(* Logix 5000 project; controller UOWHF Emulate 5570 rev 30.12; software revision 30.00; part 11 of 13 *)
(* tags used below, declared in another part *)
   UOWHF_Add_c : DINT;
   UOWHF_Msg : DINT[16];
   UOWHF_Result : DINT[16];
(* MainProgram, continued *)

   		UOWHF_Add_c.2:=UOWHF_Result[2].31;
   		UOWHF_Result[2].31:=0;
   		UOWHF_Result[3]:=UOWHF_Result[3] + 1591004397+UOWHF_Add_c;
   		UOWHF_Add_c.3:=UOWHF_Result[3].31;
   		UOWHF_Result[3].31:=0;
   		UOWHF_Result[4]:=UOWHF_Result[4] + 1640170804+UOWHF_Add_c;
   		UOWHF_Add_c.4:=UOWHF_Result[4].31;
   		UOWHF_Result[4].31:=0;
   		UOWHF_Result[5]:=UOWHF_Result[5] + 417190836+UOWHF_Add_c;
   		UOWHF_Add_c.5:=UOWHF_Result[5].31;
   		UOWHF_Result[5].31:=0;
   		UOWHF_Result[6]:=UOWHF_Result[6] + 1926019562+UOWHF_Add_c;
   		UOWHF_Add_c.6:=UOWHF_Result[6].31;
   		UOWHF_Result[6].31:=0;
   		UOWHF_Result[7]:=UOWHF_Result[7] + 695957955+UOWHF_Add_c;
   		UOWHF_Add_c.7:=UOWHF_Result[7].31;
   		UOWHF_Result[7].31:=0;
   		UOWHF_Result[8]:=UOWHF_Result[8] + 1059440084+UOWHF_Add_c;
   		UOWHF_Add_c.8:=UOWHF_Result[8].31;
   		UOWHF_Result[8].31:=0;
   	End_If;
   	If UOWHF_Msg[10].[4] Then
   		UOWHF_Result[0]:=UOWHF_Result[0] + 901796020+UOWHF_Add_c;
   		UOWHF_Add_c.0:=UOWHF_Result[0].31;
   		UOWHF_Result[0].31:=0;
   		UOWHF_Result[1]:=UOWHF_Result[1] + 1127200049+UOWHF_Add_c;
   		UOWHF_Add_c.1:=UOWHF_Result[1].31;
   		UOWHF_Result[1].31:=0;
   		UOWHF_Result[2]:=UOWHF_Result[2] + 1602413067+UOWHF_Add_c;
   		UOWHF_Add_c.2:=UOWHF_Result[2].31;
   		UOWHF_Result[2].31:=0;
   		UOWHF_Result[3]:=UOWHF_Result[3] + 1255033930+UOWHF_Add_c;
   		UOWHF_Add_c.3:=UOWHF_Result[3].31;
   		UOWHF_Result[3].31:=0;
   		UOWHF_Result[4]:=UOWHF_Result[4] + 2144327764+UOWHF_Add_c;
   		UOWHF_Add_c.4:=UOWHF_Result[4].31;
   		UOWHF_Result[4].31:=0;
   		UOWHF_Result[5]:=UOWHF_Result[5] + 1452466792+UOWHF_Add_c;
   		UOWHF_Add_c.5:=UOWHF_Result[5].31;
   		UOWHF_Result[5].31:=0;
   		UOWHF_Result[6]:=UOWHF_Result[6] + 154742090+UOWHF_Add_c;
   		UOWHF_Add_c.6:=UOWHF_Result[6].31;
   		UOWHF_Result[6].31:=0;
   		UOWHF_Result[7]:=UOWHF_Result[7] + 1902468370+UOWHF_Add_c;
   		UOWHF_Add_c.7:=UOWHF_Result[7].31;
   		UOWHF_Result[7].31:=0;
   		UOWHF_Result[8]:=UOWHF_Result[8] + 342884653+UOWHF_Add_c;
   		UOWHF_Add_c.8:=UOWHF_Result[8].31;
   		UOWHF_Result[8].31:=0;
   	End_If;
   	If UOWHF_Msg[10].[5] Then
   		UOWHF_Result[0]:=UOWHF_Result[0] + 868277617+UOWHF_Add_c;
   		UOWHF_Add_c.0:=UOWHF_Result[0].31;
   		UOWHF_Result[0].31:=0;
   		UOWHF_Result[1]:=UOWHF_Result[1] + 1436615864+UOWHF_Add_c;
   		UOWHF_Add_c.1:=UOWHF_Result[1].31;
   		UOWHF_Result[1].31:=0;
   		UOWHF_Result[2]:=UOWHF_Result[2] + 1784814025+UOWHF_Add_c;
   		UOWHF_Add_c.2:=UOWHF_Result[2].31;
   		UOWHF_Result[2].31:=0;
   		UOWHF_Result[3]:=UOWHF_Result[3] + 1380127603+UOWHF_Add_c;
   		UOWHF_Add_c.3:=UOWHF_Result[3].31;
   		UOWHF_Result[3].31:=0;
   		UOWHF_Result[4]:=UOWHF_Result[4] + 1271855125+UOWHF_Add_c;
   		UOWHF_Add_c.4:=UOWHF_Result[4].31;
   		UOWHF_Result[4].31:=0;
   		UOWHF_Result[5]:=UOWHF_Result[5] + 1937374017+UOWHF_Add_c;
   		UOWHF_Add_c.5:=UOWHF_Result[5].31;
   		UOWHF_Result[5].31:=0;
   		UOWHF_Result[6]:=UOWHF_Result[6] + 1845918423+UOWHF_Add_c;
   		UOWHF_Add_c.6:=UOWHF_Result[6].31;
   		UOWHF_Result[6].31:=0;
   		UOWHF_Result[7]:=UOWHF_Result[7] + 1463581006+UOWHF_Add_c;
   		UOWHF_Add_c.7:=UOWHF_Result[7].31;
   		UOWHF_Result[7].31:=0;
   		UOWHF_Result[8]:=UOWHF_Result[8] + 350086967+UOWHF_Add_c;
   		UOWHF_Add_c.8:=UOWHF_Result[8].31;
   		UOWHF_Result[8].31:=0;
   	End_If;
   	If UOWHF_Msg[10].[6] Then
   		UOWHF_Result[0]:=UOWHF_Result[0] + 1588271974+UOWHF_Add_c;
   		UOWHF_Add_c.0:=UOWHF_Result[0].31;
   		UOWHF_Result[0].31:=0;
   		UOWHF_Result[1]:=UOWHF_Result[1] + 586756377+UOWHF_Add_c;
   		UOWHF_Add_c.1:=UOWHF_Result[1].31;
   		UOWHF_Result[1].31:=0;
   		UOWHF_Result[2]:=UOWHF_Result[2] + 559516102+UOWHF_Add_c;
   		UOWHF_Add_c.2:=UOWHF_Result[2].31;
   		UOWHF_Result[2].31:=0;
   		UOWHF_Result[3]:=UOWHF_Result[3] + 331741523+UOWHF_Add_c;
   		UOWHF_Add_c.3:=UOWHF_Result[3].31;
   		UOWHF_Result[3].31:=0;
   		UOWHF_Result[4]:=UOWHF_Result[4] + 1880781678+UOWHF_Add_c;
   		UOWHF_Add_c.4:=UOWHF_Result[4].31;
   		UOWHF_Result[4].31:=0;
   		UOWHF_Result[5]:=UOWHF_Result[5] + 1152892566+UOWHF_Add_c;
   		UOWHF_Add_c.5:=UOWHF_Result[5].31;
   		UOWHF_Result[5].31:=0;
   		UOWHF_Result[6]:=UOWHF_Result[6] + 2047233698+UOWHF_Add_c;
   		UOWHF_Add_c.6:=UOWHF_Result[6].31;
   		UOWHF_Result[6].31:=0;
   		UOWHF_Result[7]:=UOWHF_Result[7] + 1642594289+UOWHF_Add_c;
   		UOWHF_Add_c.7:=UOWHF_Result[7].31;
   		UOWHF_Result[7].31:=0;
   		UOWHF_Result[8]:=UOWHF_Result[8] + 376585573+UOWHF_Add_c;
   		UOWHF_Add_c.8:=UOWHF_Result[8].31;
   		UOWHF_Result[8].31:=0;
   	End_If;
   	If UOWHF_Msg[10].[7] Then
   		UOWHF_Result[0]:=UOWHF_Result[0] + 1020715491+UOWHF_Add_c;
   		UOWHF_Add_c.0:=UOWHF_Result[0].31;
   		UOWHF_Result[0].31:=0;
   		UOWHF_Result[1]:=UOWHF_Result[1] + 1857205629+UOWHF_Add_c;
   		UOWHF_Add_c.1:=UOWHF_Result[1].31;
   		UOWHF_Result[1].31:=0;
   		UOWHF_Result[2]:=UOWHF_Result[2] + 16853309+UOWHF_Add_c;
   		UOWHF_Add_c.2:=UOWHF_Result[2].31;
   		UOWHF_Result[2].31:=0;
   		UOWHF_Result[3]:=UOWHF_Result[3] + 1231994168+UOWHF_Add_c;
   		UOWHF_Add_c.3:=UOWHF_Result[3].31;
   		UOWHF_Result[3].31:=0;
   		UOWHF_Result[4]:=UOWHF_Result[4] + 423998966+UOWHF_Add_c;
   		UOWHF_Add_c.4:=UOWHF_Result[4].31;
   		UOWHF_Result[4].31:=0;
   		UOWHF_Result[5]:=UOWHF_Result[5] + 1299862752+UOWHF_Add_c;
   		UOWHF_Add_c.5:=UOWHF_Result[5].31;
   		UOWHF_Result[5].31:=0;
   		UOWHF_Result[6]:=UOWHF_Result[6] + 652509862+UOWHF_Add_c;
   		UOWHF_Add_c.6:=UOWHF_Result[6].31;
   		UOWHF_Result[6].31:=0;
   		UOWHF_Result[7]:=UOWHF_Result[7] + 15353685+UOWHF_Add_c;
   		UOWHF_Add_c.7:=UOWHF_Result[7].31;
   		UOWHF_Result[7].31:=0;
   		UOWHF_Result[8]:=UOWHF_Result[8] + 2001428660+UOWHF_Add_c;
   		UOWHF_Add_c.8:=UOWHF_Result[8].31;
   		UOWHF_Result[8].31:=0;
   	End_If;
   	If UOWHF_Msg[10].[8] Then
   		UOWHF_Result[0]:=UOWHF_Result[0] + 813810484+UOWHF_Add_c;
   		UOWHF_Add_c.0:=UOWHF_Result[0].31;
   		UOWHF_Result[0].31:=0;
   		UOWHF_Result[1]:=UOWHF_Result[1] + 1003989381+UOWHF_Add_c;
   		UOWHF_Add_c.1:=UOWHF_Result[1].31;
   		UOWHF_Result[1].31:=0;
   		UOWHF_Result[2]:=UOWHF_Result[2] + 738018774+UOWHF_Add_c;
   		UOWHF_Add_c.2:=UOWHF_Result[2].31;
   		UOWHF_Result[2].31:=0;
   		UOWHF_Result[3]:=UOWHF_Result[3] + 443461312+UOWHF_Add_c;
   		UOWHF_Add_c.3:=UOWHF_Result[3].31;
   		UOWHF_Result[3].31:=0;
   		UOWHF_Result[4]:=UOWHF_Result[4] + 1637414295+UOWHF_Add_c;
   		UOWHF_Add_c.4:=UOWHF_Result[4].31;
   		UOWHF_Result[4].31:=0;
   		UOWHF_Result[5]:=UOWHF_Result[5] + 157939787+UOWHF_Add_c;
   		UOWHF_Add_c.5:=UOWHF_Result[5].31;
   		UOWHF_Result[5].31:=0;
   		UOWHF_Result[6]:=UOWHF_Result[6] + 712235666+UOWHF_Add_c;
   		UOWHF_Add_c.6:=UOWHF_Result[6].31;
   		UOWHF_Result[6].31:=0;
   		UOWHF_Result[7]:=UOWHF_Result[7] + 1688386276+UOWHF_Add_c;
   		UOWHF_Add_c.7:=UOWHF_Result[7].31;
   		UOWHF_Result[7].31:=0;
   		UOWHF_Result[8]:=UOWHF_Result[8] + 2013177678+UOWHF_Add_c;
   		UOWHF_Add_c.8:=UOWHF_Result[8].31;
   		UOWHF_Result[8].31:=0;
   	End_If;
   	If UOWHF_Msg[10].[9] Then
   		UOWHF_Result[0]:=UOWHF_Result[0] + 1535414445+UOWHF_Add_c;
   		UOWHF_Add_c.0:=UOWHF_Result[0].31;
   		UOWHF_Result[0].31:=0;
   		UOWHF_Result[1]:=UOWHF_Result[1] + 1615623515+UOWHF_Add_c;
   		UOWHF_Add_c.1:=UOWHF_Result[1].31;
   		UOWHF_Result[1].31:=0;
   		UOWHF_Result[2]:=UOWHF_Result[2] + 1360597756+UOWHF_Add_c;
   		UOWHF_Add_c.2:=UOWHF_Result[2].31;
   		UOWHF_Result[2].31:=0;
   		UOWHF_Result[3]:=UOWHF_Result[3] + 1573823097+UOWHF_Add_c;
   		UOWHF_Add_c.3:=UOWHF_Result[3].31;
   		UOWHF_Result[3].31:=0;
   		UOWHF_Result[4]:=UOWHF_Result[4] + 1281710714+UOWHF_Add_c;
   		UOWHF_Add_c.4:=UOWHF_Result[4].31;
   		UOWHF_Result[4].31:=0;
   		UOWHF_Result[5]:=UOWHF_Result[5] + 1453733315+UOWHF_Add_c;
   		UOWHF_Add_c.5:=UOWHF_Result[5].31;
   		UOWHF_Result[5].31:=0;
   		UOWHF_Result[6]:=UOWHF_Result[6] + 369997754+UOWHF_Add_c;
   		UOWHF_Add_c.6:=UOWHF_Result[6].31;
   		UOWHF_Result[6].31:=0;
   		UOWHF_Result[7]:=UOWHF_Result[7] + 1856281529+UOWHF_Add_c;
   		UOWHF_Add_c.7:=UOWHF_Result[7].31;
   		UOWHF_Result[7].31:=0;
   		UOWHF_Result[8]:=UOWHF_Result[8] + 1847238559+UOWHF_Add_c;
   		UOWHF_Add_c.8:=UOWHF_Result[8].31;
   		UOWHF_Result[8].31:=0;
   	End_If;
   	If UOWHF_Msg[10].[10] Then
   		UOWHF_Result[0]:=UOWHF_Result[0] + 1061749827+UOWHF_Add_c;
   		UOWHF_Add_c.0:=UOWHF_Result[0].31;
   		UOWHF_Result[0].31:=0;
   		UOWHF_Result[1]:=UOWHF_Result[1] + 842932244+UOWHF_Add_c;
   		UOWHF_Add_c.1:=UOWHF_Result[1].31;
   		UOWHF_Result[1].31:=0;
   		UOWHF_Result[2]:=UOWHF_Result[2] + 1033461891+UOWHF_Add_c;
   		UOWHF_Add_c.2:=UOWHF_Result[2].31;
   		UOWHF_Result[2].31:=0;
   		UOWHF_Result[3]:=UOWHF_Result[3] + 379746348+UOWHF_Add_c;
   		UOWHF_Add_c.3:=UOWHF_Result[3].31;
   		UOWHF_Result[3].31:=0;
   		UOWHF_Result[4]:=UOWHF_Result[4] + 685495130+UOWHF_Add_c;
   		UOWHF_Add_c.4:=UOWHF_Result[4].31;
   		UOWHF_Result[4].31:=0;
   		UOWHF_Result[5]:=UOWHF_Result[5] + 958802377+UOWHF_Add_c;
   		UOWHF_Add_c.5:=UOWHF_Result[5].31;
   		UOWHF_Result[5].31:=0;
   		UOWHF_Result[6]:=UOWHF_Result[6] + 129067151+UOWHF_Add_c;
   		UOWHF_Add_c.6:=UOWHF_Result[6].31;
   		UOWHF_Result[6].31:=0;
   		UOWHF_Result[7]:=UOWHF_Result[7] + 1694766568+UOWHF_Add_c;
   		UOWHF_Add_c.7:=UOWHF_Result[7].31;
   		UOWHF_Result[7].31:=0;
   		UOWHF_Result[8]:=UOWHF_Result[8] + 1431412769+UOWHF_Add_c;
   		UOWHF_Add_c.8:=UOWHF_Result[8].31;
   		UOWHF_Result[8].31:=0;
   	End_If;
   	If UOWHF_Msg[10].[11] Then
   		UOWHF_Result[0]:=UOWHF_Result[0] + 1646350318+UOWHF_Add_c;
   		UOWHF_Add_c.0:=UOWHF_Result[0].31;
   		UOWHF_Result[0].31:=0;
   		UOWHF_Result[1]:=UOWHF_Result[1] + 1974652699+UOWHF_Add_c;
   		UOWHF_Add_c.1:=UOWHF_Result[1].31;
   		UOWHF_Result[1].31:=0;
   		UOWHF_Result[2]:=UOWHF_Result[2] + 325775484+UOWHF_Add_c;
   		UOWHF_Add_c.2:=UOWHF_Result[2].31;
   		UOWHF_Result[2].31:=0;
   		UOWHF_Result[3]:=UOWHF_Result[3] + 83362006+UOWHF_Add_c;
   		UOWHF_Add_c.3:=UOWHF_Result[3].31;
   		UOWHF_Result[3].31:=0;
   		UOWHF_Result[4]:=UOWHF_Result[4] + 262049431+UOWHF_Add_c;
   		UOWHF_Add_c.4:=UOWHF_Result[4].31;
   		UOWHF_Result[4].31:=0;
   		UOWHF_Result[5]:=UOWHF_Result[5] + 1644755762+UOWHF_Add_c;
   		UOWHF_Add_c.5:=UOWHF_Result[5].31;
   		UOWHF_Result[5].31:=0;
   		UOWHF_Result[6]:=UOWHF_Result[6] + 790241358+UOWHF_Add_c;
   		UOWHF_Add_c.6:=UOWHF_Result[6].31;
   		UOWHF_Result[6].31:=0;
   		UOWHF_Result[7]:=UOWHF_Result[7] + 2126439262+UOWHF_Add_c;
   		UOWHF_Add_c.7:=UOWHF_Result[7].31;
   		UOWHF_Result[7].31:=0;
   		UOWHF_Result[8]:=UOWHF_Result[8] + 1052212769+UOWHF_Add_c;
   		UOWHF_Add_c.8:=UOWHF_Result[8].31;
   		UOWHF_Result[8].31:=0;
   	End_If;
   	If UOWHF_Msg[10].[12] Then
   		UOWHF_Result[0]:=UOWHF_Result[0] + 955937059+UOWHF_Add_c;
   		UOWHF_Add_c.0:=UOWHF_Result[0].31;
   		UOWHF_Result[0].31:=0;
   		UOWHF_Result[1]:=UOWHF_Result[1] + 936365642+UOWHF_Add_c;
   		UOWHF_Add_c.1:=UOWHF_Result[1].31;
   		UOWHF_Result[1].31:=0;
   		UOWHF_Result[2]:=UOWHF_Result[2] + 498042732+UOWHF_Add_c;
   		UOWHF_Add_c.2:=UOWHF_Result[2].31;
   		UOWHF_Result[2].31:=0;
   		UOWHF_Result[3]:=UOWHF_Result[3] + 238009702+UOWHF_Add_c;
   		UOWHF_Add_c.3:=UOWHF_Result[3].31;
   		UOWHF_Result[3].31:=0;
   		UOWHF_Result[4]:=UOWHF_Result[4] + 36957456+UOWHF_Add_c;
   		UOWHF_Add_c.4:=UOWHF_Result[4].31;
   		UOWHF_Result[4].31:=0;
   		UOWHF_Result[5]:=UOWHF_Result[5] + 598813011+UOWHF_Add_c;
   		UOWHF_Add_c.5:=UOWHF_Result[5].31;
   		UOWHF_Result[5].31:=0;
   		UOWHF_Result[6]:=UOWHF_Result[6] + 426350274+UOWHF_Add_c;
   		UOWHF_Add_c.6:=UOWHF_Result[6].31;
   		UOWHF_Result[6].31:=0;
   		UOWHF_Result[7]:=UOWHF_Result[7] + 102852187+UOWHF_Add_c;
   		UOWHF_Add_c.7:=UOWHF_Result[7].31;
   		UOWHF_Result[7].31:=0;
   		UOWHF_Result[8]:=UOWHF_Result[8] + 1154127904+UOWHF_Add_c;
   		UOWHF_Add_c.8:=UOWHF_Result[8].31;
   		UOWHF_Result[8].31:=0;
   	End_If;
   	If UOWHF_Msg[10].[13] Then
   		UOWHF_Result[0]:=UOWHF_Result[0] + 1268816444+UOWHF_Add_c;
   		UOWHF_Add_c.0:=UOWHF_Result[0].31;
   		UOWHF_Result[0].31:=0;
   		UOWHF_Result[1]:=UOWHF_Result[1] + 1033144398+UOWHF_Add_c;
   		UOWHF_Add_c.1:=UOWHF_Result[1].31;
   		UOWHF_Result[1].31:=0;
   		UOWHF_Result[2]:=UOWHF_Result[2] + 2027448386+UOWHF_Add_c;
   		UOWHF_Add_c.2:=UOWHF_Result[2].31;
   		UOWHF_Result[2].31:=0;
   		UOWHF_Result[3]:=UOWHF_Result[3] + 885764043+UOWHF_Add_c;
   		UOWHF_Add_c.3:=UOWHF_Result[3].31;
   		UOWHF_Result[3].31:=0;
   		UOWHF_Result[4]:=UOWHF_Result[4] + 1657422268+UOWHF_Add_c;
   		UOWHF_Add_c.4:=UOWHF_Result[4].31;
   		UOWHF_Result[4].31:=0;
   		UOWHF_Result[5]:=UOWHF_Result[5] + 1988850223+UOWHF_Add_c;
   		UOWHF_Add_c.5:=UOWHF_Result[5].31;
   		UOWHF_Result[5].31:=0;
   		UOWHF_Result[6]:=UOWHF_Result[6] + 1530930092+UOWHF_Add_c;
   		UOWHF_Add_c.6:=UOWHF_Result[6].31;
   		UOWHF_Result[6].31:=0;
   		UOWHF_Result[7]:=UOWHF_Result[7] + 2006297248+UOWHF_Add_c;
   		UOWHF_Add_c.7:=UOWHF_Result[7].31;
   		UOWHF_Result[7].31:=0;
   		UOWHF_Result[8]:=UOWHF_Result[8] + 2077959681+UOWHF_Add_c;
   		UOWHF_Add_c.8:=UOWHF_Result[8].31;
   		UOWHF_Result[8].31:=0;
   	End_If;
   	If UOWHF_Msg[10].[14] Then
   		UOWHF_Result[0]:=UOWHF_Result[0] + 1110917864+UOWHF_Add_c;
   		UOWHF_Add_c.0:=UOWHF_Result[0].31;
   		UOWHF_Result[0].31:=0;
   		UOWHF_Result[1]:=UOWHF_Result[1] + 1451124381+UOWHF_Add_c;
   		UOWHF_Add_c.1:=UOWHF_Result[1].31;
   		UOWHF_Result[1].31:=0;
   		UOWHF_Result[2]:=UOWHF_Result[2] + 1354761017+UOWHF_Add_c;
   		UOWHF_Add_c.2:=UOWHF_Result[2].31;
   		UOWHF_Result[2].31:=0;
   		UOWHF_Result[3]:=UOWHF_Result[3] + 38190742+UOWHF_Add_c;
   		UOWHF_Add_c.3:=UOWHF_Result[3].31;
   		UOWHF_Result[3].31:=0;
   		UOWHF_Result[4]:=UOWHF_Result[4] + 1921805953+UOWHF_Add_c;
   		UOWHF_Add_c.4:=UOWHF_Result[4].31;
   		UOWHF_Result[4].31:=0;
   		UOWHF_Result[5]:=UOWHF_Result[5] + 1941105002+UOWHF_Add_c;
   		UOWHF_Add_c.5:=UOWHF_Result[5].31;
   		UOWHF_Result[5].31:=0;
   		UOWHF_Result[6]:=UOWHF_Result[6] + 1703548468+UOWHF_Add_c;
   		UOWHF_Add_c.6:=UOWHF_Result[6].31;
   		UOWHF_Result[6].31:=0;
   		UOWHF_Result[7]:=UOWHF_Result[7] + 186991094+UOWHF_Add_c;
   		UOWHF_Add_c.7:=UOWHF_Result[7].31;
   		UOWHF_Result[7].31:=0;
   		UOWHF_Result[8]:=UOWHF_Result[8] + 714064657+UOWHF_Add_c;
   		UOWHF_Add_c.8:=UOWHF_Result[8].31;
   		UOWHF_Result[8].31:=0;
   	End_If;
   	If UOWHF_Msg[10].[15] Then
   		UOWHF_Result[0]:=UOWHF_Result[0] + 1961147110+UOWHF_Add_c;
   		UOWHF_Add_c.0:=UOWHF_Result[0].31;
   		UOWHF_Result[0].31:=0;
   		UOWHF_Result[1]:=UOWHF_Result[1] + 12565547+UOWHF_Add_c;
   		UOWHF_Add_c.1:=UOWHF_Result[1].31;
   		UOWHF_Result[1].31:=0;
   		UOWHF_Result[2]:=UOWHF_Result[2] + 567043951+UOWHF_Add_c;
   		UOWHF_Add_c.2:=UOWHF_Result[2].31;
   		UOWHF_Result[2].31:=0;
   		UOWHF_Result[3]:=UOWHF_Result[3] + 65949662+UOWHF_Add_c;
   		UOWHF_Add_c.3:=UOWHF_Result[3].31;
   		UOWHF_Result[3].31:=0;
   		UOWHF_Result[4]:=UOWHF_Result[4] + 1646539206+UOWHF_Add_c;
   		UOWHF_Add_c.4:=UOWHF_Result[4].31;
   		UOWHF_Result[4].31:=0;
   		UOWHF_Result[5]:=UOWHF_Result[5] + 1708716662+UOWHF_Add_c;
   		UOWHF_Add_c.5:=UOWHF_Result[5].31;
   		UOWHF_Result[5].31:=0;
   		UOWHF_Result[6]:=UOWHF_Result[6] + 1848936862+UOWHF_Add_c;
   		UOWHF_Add_c.6:=UOWHF_Result[6].31;
   		UOWHF_Result[6].31:=0;
   		UOWHF_Result[7]:=UOWHF_Result[7] + 1900654345+UOWHF_Add_c;
   		UOWHF_Add_c.7:=UOWHF_Result[7].31;
   		UOWHF_Result[7].31:=0;
   		UOWHF_Result[8]:=UOWHF_Result[8] + 1004361316+UOWHF_Add_c;
   		UOWHF_Add_c.8:=UOWHF_Result[8].31;
   		UOWHF_Result[8].31:=0;
   	End_If;
   	If UOWHF_Msg[10].[16] Then
   		UOWHF_Result[0]:=UOWHF_Result[0] + 415520432+UOWHF_Add_c;
   		UOWHF_Add_c.0:=UOWHF_Result[0].31;
   		UOWHF_Result[0].31:=0;
   		UOWHF_Result[1]:=UOWHF_Result[1] + 351467464+UOWHF_Add_c;
   		UOWHF_Add_c.1:=UOWHF_Result[1].31;
   		UOWHF_Result[1].31:=0;
   		UOWHF_Result[2]:=UOWHF_Result[2] + 654166220+UOWHF_Add_c;
   		UOWHF_Add_c.2:=UOWHF_Result[2].31;
   		UOWHF_Result[2].31:=0;
   		UOWHF_Result[3]:=UOWHF_Result[3] + 741029837+UOWHF_Add_c;
   		UOWHF_Add_c.3:=UOWHF_Result[3].31;
   		UOWHF_Result[3].31:=0;
   		UOWHF_Result[4]:=UOWHF_Result[4] + 1981690344+UOWHF_Add_c;
   		UOWHF_Add_c.4:=UOWHF_Result[4].31;
   		UOWHF_Result[4].31:=0;
   		UOWHF_Result[5]:=UOWHF_Result[5] + 19210638+UOWHF_Add_c;
   		UOWHF_Add_c.5:=UOWHF_Result[5].31;
   		UOWHF_Result[5].31:=0;
   		UOWHF_Result[6]:=UOWHF_Result[6] + 566229794+UOWHF_Add_c;
   		UOWHF_Add_c.6:=UOWHF_Result[6].31;
   		UOWHF_Result[6].31:=0;
   		UOWHF_Result[7]:=UOWHF_Result[7] + 625793338+UOWHF_Add_c;
   		UOWHF_Add_c.7:=UOWHF_Result[7].31;
   		UOWHF_Result[7].31:=0;
   		UOWHF_Result[8]:=UOWHF_Result[8] + 386405378+UOWHF_Add_c;
   		UOWHF_Add_c.8:=UOWHF_Result[8].31;
   		UOWHF_Result[8].31:=0;
   	End_If;
   	If UOWHF_Msg[10].[17] Then
   		UOWHF_Result[0]:=UOWHF_Result[0] + 1499883797+UOWHF_Add_c;
   		UOWHF_Add_c.0:=UOWHF_Result[0].31;
   		UOWHF_Result[0].31:=0;
   		UOWHF_Result[1]:=UOWHF_Result[1] + 129680376+UOWHF_Add_c;
   		UOWHF_Add_c.1:=UOWHF_Result[1].31;
   		UOWHF_Result[1].31:=0;
   		UOWHF_Result[2]:=UOWHF_Result[2] + 700971919+UOWHF_Add_c;
   		UOWHF_Add_c.2:=UOWHF_Result[2].31;
   		UOWHF_Result[2].31:=0;
   		UOWHF_Result[3]:=UOWHF_Result[3] + 56395807+UOWHF_Add_c;
   		UOWHF_Add_c.3:=UOWHF_Result[3].31;
   		UOWHF_Result[3].31:=0;
   		UOWHF_Result[4]:=UOWHF_Result[4] + 1355965327+UOWHF_Add_c;
   		UOWHF_Add_c.4:=UOWHF_Result[4].31;
   		UOWHF_Result[4].31:=0;
   		UOWHF_Result[5]:=UOWHF_Result[5] + 1408183226+UOWHF_Add_c;
   		UOWHF_Add_c.5:=UOWHF_Result[5].31;
   		UOWHF_Result[5].31:=0;
   		UOWHF_Result[6]:=UOWHF_Result[6] + 2071090026+UOWHF_Add_c;
   		UOWHF_Add_c.6:=UOWHF_Result[6].31;
   		UOWHF_Result[6].31:=0;
   		UOWHF_Result[7]:=UOWHF_Result[7] + 1334749712+UOWHF_Add_c;
   		UOWHF_Add_c.7:=UOWHF_Result[7].31;
   		UOWHF_Result[7].31:=0;
   		UOWHF_Result[8]:=UOWHF_Result[8] + 894206129+UOWHF_Add_c;
   		UOWHF_Add_c.8:=UOWHF_Result[8].31;
   		UOWHF_Result[8].31:=0;
   	End_If;
   	If UOWHF_Msg[10].[18] Then
   		UOWHF_Result[0]:=UOWHF_Result[0] + 611633887+UOWHF_Add_c;
   		UOWHF_Add_c.0:=UOWHF_Result[0].31;
   		UOWHF_Result[0].31:=0;
   		UOWHF_Result[1]:=UOWHF_Result[1] + 220479088+UOWHF_Add_c;
   		UOWHF_Add_c.1:=UOWHF_Result[1].31;
   		UOWHF_Result[1].31:=0;
   		UOWHF_Result[2]:=UOWHF_Result[2] + 774163886+UOWHF_Add_c;
   		UOWHF_Add_c.2:=UOWHF_Result[2].31;
   		UOWHF_Result[2].31:=0;
   		UOWHF_Result[3]:=UOWHF_Result[3] + 244973967+UOWHF_Add_c;
   		UOWHF_Add_c.3:=UOWHF_Result[3].31;
   		UOWHF_Result[3].31:=0;
   		UOWHF_Result[4]:=UOWHF_Result[4] + 906891116+UOWHF_Add_c;
   		UOWHF_Add_c.4:=UOWHF_Result[4].31;
   		UOWHF_Result[4].31:=0;
   		UOWHF_Result[5]:=UOWHF_Result[5] + 2010017338+UOWHF_Add_c;
   		UOWHF_Add_c.5:=UOWHF_Result[5].31;
   		UOWHF_Result[5].31:=0;
   		UOWHF_Result[6]:=UOWHF_Result[6] + 1437360572+UOWHF_Add_c;
   		UOWHF_Add_c.6:=UOWHF_Result[6].31;
   		UOWHF_Result[6].31:=0;
   		UOWHF_Result[7]:=UOWHF_Result[7] + 1208873370+UOWHF_Add_c;
   		UOWHF_Add_c.7:=UOWHF_Result[7].31;
   		UOWHF_Result[7].31:=0;
   		UOWHF_Result[8]:=UOWHF_Result[8] + 73161532+UOWHF_Add_c;
   		UOWHF_Add_c.8:=UOWHF_Result[8].31;
   		UOWHF_Result[8].31:=0;
   	End_If;
   	If UOWHF_Msg[10].[19] Then
   		UOWHF_Result[0]:=UOWHF_Result[0] + 1276434743+UOWHF_Add_c;
   		UOWHF_Add_c.0:=UOWHF_Result[0].31;
   		UOWHF_Result[0].31:=0;
   		UOWHF_Result[1]:=UOWHF_Result[1] + 923954815+UOWHF_Add_c;
   		UOWHF_Add_c.1:=UOWHF_Result[1].31;
   		UOWHF_Result[1].31:=0;
   		UOWHF_Result[2]:=UOWHF_Result[2] + 2127328610+UOWHF_Add_c;
   		UOWHF_Add_c.2:=UOWHF_Result[2].31;
   		UOWHF_Result[2].31:=0;
   		UOWHF_Result[3]:=UOWHF_Result[3] + 1862713612+UOWHF_Add_c;
   		UOWHF_Add_c.3:=UOWHF_Result[3].31;
   		UOWHF_Result[3].31:=0;
   		UOWHF_Result[4]:=UOWHF_Result[4] + 1878938249+UOWHF_Add_c;
   		UOWHF_Add_c.4:=UOWHF_Result[4].31;
   		UOWHF_Result[4].31:=0;
   		UOWHF_Result[5]:=UOWHF_Result[5] + 1189510329+UOWHF_Add_c;
   		UOWHF_Add_c.5:=UOWHF_Result[5].31;
   		UOWHF_Result[5].31:=0;
   		UOWHF_Result[6]:=UOWHF_Result[6] + 1679535384+UOWHF_Add_c;
   		UOWHF_Add_c.6:=UOWHF_Result[6].31;
   		UOWHF_Result[6].31:=0;
   		UOWHF_Result[7]:=UOWHF_Result[7] + 1749990172+UOWHF_Add_c;
   		UOWHF_Add_c.7:=UOWHF_Result[7].31;
   		UOWHF_Result[7].31:=0;
   		UOWHF_Result[8]:=UOWHF_Result[8] + 1880399620+UOWHF_Add_c;
   		UOWHF_Add_c.8:=UOWHF_Result[8].31;
   		UOWHF_Result[8].31:=0;
   	End_If;
   	If UOWHF_Msg[10].[20] Then
   		UOWHF_Result[0]:=UOWHF_Result[0] + 1067539284+UOWHF_Add_c;
   		UOWHF_Add_c.0:=UOWHF_Result[0].31;
   		UOWHF_Result[0].31:=0;
   		UOWHF_Result[1]:=UOWHF_Result[1] + 1218546281+UOWHF_Add_c;
   		UOWHF_Add_c.1:=UOWHF_Result[1].31;
   		UOWHF_Result[1].31:=0;
   		UOWHF_Result[2]:=UOWHF_Result[2] + 1692266167+UOWHF_Add_c;
   		UOWHF_Add_c.2:=UOWHF_Result[2].31;
   		UOWHF_Result[2].31:=0;
   		UOWHF_Result[3]:=UOWHF_Result[3] + 844450602+UOWHF_Add_c;
   		UOWHF_Add_c.3:=UOWHF_Result[3].31;
   		UOWHF_Result[3].31:=0;
   		UOWHF_Result[4]:=UOWHF_Result[4] + 1351238461+UOWHF_Add_c;
   		UOWHF_Add_c.4:=UOWHF_Result[4].31;
   		UOWHF_Result[4].31:=0;
   		UOWHF_Result[5]:=UOWHF_Result[5] + 2074939840+UOWHF_Add_c;
   		UOWHF_Add_c.5:=UOWHF_Result[5].31;
   		UOWHF_Result[5].31:=0;
   		UOWHF_Result[6]:=UOWHF_Result[6] + 54095456+UOWHF_Add_c;
   		UOWHF_Add_c.6:=UOWHF_Result[6].31;
   		UOWHF_Result[6].31:=0;
   		UOWHF_Result[7]:=UOWHF_Result[7] + 1472659390+UOWHF_Add_c;
   		UOWHF_Add_c.7:=UOWHF_Result[7].31;
   		UOWHF_Result[7].31:=0;
   		UOWHF_Result[8]:=UOWHF_Result[8] + 78847011+UOWHF_Add_c;
   		UOWHF_Add_c.8:=UOWHF_Result[8].31;
   		UOWHF_Result[8].31:=0;
   	End_If;
   	If UOWHF_Msg[10].[21] Then
   		UOWHF_Result[0]:=UOWHF_Result[0] + 615459290+UOWHF_Add_c;
   		UOWHF_Add_c.0:=UOWHF_Result[0].31;
   		UOWHF_Result[0].31:=0;
   		UOWHF_Result[1]:=UOWHF_Result[1] + 628300652+UOWHF_Add_c;
   		UOWHF_Add_c.1:=UOWHF_Result[1].31;
   		UOWHF_Result[1].31:=0;
   		UOWHF_Result[2]:=UOWHF_Result[2] + 913630562+UOWHF_Add_c;
   		UOWHF_Add_c.2:=UOWHF_Result[2].31;
   		UOWHF_Result[2].31:=0;
   		UOWHF_Result[3]:=UOWHF_Result[3] + 1573973421+UOWHF_Add_c;
   		UOWHF_Add_c.3:=UOWHF_Result[3].31;
   		UOWHF_Result[3].31:=0;
   		UOWHF_Result[4]:=UOWHF_Result[4] + 842720559+UOWHF_Add_c;
   		UOWHF_Add_c.4:=UOWHF_Result[4].31;
   		UOWHF_Result[4].31:=0;
   		UOWHF_Result[5]:=UOWHF_Result[5] + 1465717949+UOWHF_Add_c;
   		UOWHF_Add_c.5:=UOWHF_Result[5].31;
   		UOWHF_Result[5].31:=0;
   		UOWHF_Result[6]:=UOWHF_Result[6] + 1475649611+UOWHF_Add_c;
   		UOWHF_Add_c.6:=UOWHF_Result[6].31;
   		UOWHF_Result[6].31:=0;
   		UOWHF_Result[7]:=UOWHF_Result[7] + 1123747716+UOWHF_Add_c;
   		UOWHF_Add_c.7:=UOWHF_Result[7].31;
   		UOWHF_Result[7].31:=0;
   		UOWHF_Result[8]:=UOWHF_Result[8] + 593611670+UOWHF_Add_c;
   		UOWHF_Add_c.8:=UOWHF_Result[8].31;
   		UOWHF_Result[8].31:=0;
   	End_If;
   	If UOWHF_Msg[10].[22] Then
   		UOWHF_Result[0]:=UOWHF_Result[0] + 333024015+UOWHF_Add_c;
   		UOWHF_Add_c.0:=UOWHF_Result[0].31;
   		UOWHF_Result[0].31:=0;
   		UOWHF_Result[1]:=UOWHF_Result[1] + 649171931+UOWHF_Add_c;
   		UOWHF_Add_c.1:=UOWHF_Result[1].31;
   		UOWHF_Result[1].31:=0;
   		UOWHF_Result[2]:=UOWHF_Result[2] + 1523497291+UOWHF_Add_c;
   		UOWHF_Add_c.2:=UOWHF_Result[2].31;
   		UOWHF_Result[2].31:=0;
   		UOWHF_Result[3]:=UOWHF_Result[3] + 1354970453+UOWHF_Add_c;
   		UOWHF_Add_c.3:=UOWHF_Result[3].31;
   		UOWHF_Result[3].31:=0;
   		UOWHF_Result[4]:=UOWHF_Result[4] + 72262000+UOWHF_Add_c;
   		UOWHF_Add_c.4:=UOWHF_Result[4].31;
   		UOWHF_Result[4].31:=0;
   		UOWHF_Result[5]:=UOWHF_Result[5] + 246209462+UOWHF_Add_c;
   		UOWHF_Add_c.5:=UOWHF_Result[5].31;
   		UOWHF_Result[5].31:=0;
   		UOWHF_Result[6]:=UOWHF_Result[6] + 1497013496+UOWHF_Add_c;
   		UOWHF_Add_c.6:=UOWHF_Result[6].31;
   		UOWHF_Result[6].31:=0;
   		UOWHF_Result[7]:=UOWHF_Result[7] + 133031163+UOWHF_Add_c;
   		UOWHF_Add_c.7:=UOWHF_Result[7].31;
   		UOWHF_Result[7].31:=0;
   		UOWHF_Result[8]:=UOWHF_Result[8] + 1209415317+UOWHF_Add_c;
   		UOWHF_Add_c.8:=UOWHF_Result[8].31;
   		UOWHF_Result[8].31:=0;
   	End_If;
   	If UOWHF_Msg[10].[23] Then
   		UOWHF_Result[0]:=UOWHF_Result[0] + 1058819959+UOWHF_Add_c;
   		UOWHF_Add_c.0:=UOWHF_Result[0].31;
   		UOWHF_Result[0].31:=0;
   		UOWHF_Result[1]:=UOWHF_Result[1] + 1490152365+UOWHF_Add_c;
   		UOWHF_Add_c.1:=UOWHF_Result[1].31;
   		UOWHF_Result[1].31:=0;
   		UOWHF_Result[2]:=UOWHF_Result[2] + 750844208+UOWHF_Add_c;
   		UOWHF_Add_c.2:=UOWHF_Result[2].31;
   		UOWHF_Result[2].31:=0;
   		UOWHF_Result[3]:=UOWHF_Result[3] + 69060592+UOWHF_Add_c;
   		UOWHF_Add_c.3:=UOWHF_Result[3].31;
   		UOWHF_Result[3].31:=0;
   		UOWHF_Result[4]:=UOWHF_Result[4] + 1239135017+UOWHF_Add_c;
   		UOWHF_Add_c.4:=UOWHF_Result[4].31;
   		UOWHF_Result[4].31:=0;
   		UOWHF_Result[5]:=UOWHF_Result[5] + 1324052255+UOWHF_Add_c;
   		UOWHF_Add_c.5:=UOWHF_Result[5].31;
   		UOWHF_Result[5].31:=0;
   		UOWHF_Result[6]:=UOWHF_Result[6] + 464992231+UOWHF_Add_c;
   		UOWHF_Add_c.6:=UOWHF_Result[6].31;
   		UOWHF_Result[6].31:=0;
   		UOWHF_Result[7]:=UOWHF_Result[7] + 903984470+UOWHF_Add_c;
   		UOWHF_Add_c.7:=UOWHF_Result[7].31;
   		UOWHF_Result[7].31:=0;
   		UOWHF_Result[8]:=UOWHF_Result[8] + 493288648+UOWHF_Add_c;
   		UOWHF_Add_c.8:=UOWHF_Result[8].31;
   		UOWHF_Result[8].31:=0;
   	End_If;
   	If UOWHF_Msg[10].[24] Then
   		UOWHF_Result[0]:=UOWHF_Result[0] + 2042370017+UOWHF_Add_c;
   		UOWHF_Add_c.0:=UOWHF_Result[0].31;
   		UOWHF_Result[0].31:=0;
   		UOWHF_Result[1]:=UOWHF_Result[1] + 499230009+UOWHF_Add_c;
   		UOWHF_Add_c.1:=UOWHF_Result[1].31;
   		UOWHF_Result[1].31:=0;
   		UOWHF_Result[2]:=UOWHF_Result[2] + 897236454+UOWHF_Add_c;
   		UOWHF_Add_c.2:=UOWHF_Result[2].31;
   		UOWHF_Result[2].31:=0;
   		UOWHF_Result[3]:=UOWHF_Result[3] + 1564035470+UOWHF_Add_c;
   		UOWHF_Add_c.3:=UOWHF_Result[3].31;
   		UOWHF_Result[3].31:=0;
   		UOWHF_Result[4]:=UOWHF_Result[4] + 1571293463+UOWHF_Add_c;
   		UOWHF_Add_c.4:=UOWHF_Result[4].31;
   		UOWHF_Result[4].31:=0;
   		UOWHF_Result[5]:=UOWHF_Result[5] + 1430387324+UOWHF_Add_c;
   		UOWHF_Add_c.5:=UOWHF_Result[5].31;
   		UOWHF_Result[5].31:=0;
   		UOWHF_Result[6]:=UOWHF_Result[6] + 468146450+UOWHF_Add_c;
   		UOWHF_Add_c.6:=UOWHF_Result[6].31;
   		UOWHF_Result[6].31:=0;
   		UOWHF_Result[7]:=UOWHF_Result[7] + 974707670+UOWHF_Add_c;
   		UOWHF_Add_c.7:=UOWHF_Result[7].31;
   		UOWHF_Result[7].31:=0;
   		UOWHF_Result[8]:=UOWHF_Result[8] + 1284040803+UOWHF_Add_c;
   		UOWHF_Add_c.8:=UOWHF_Result[8].31;
   		UOWHF_Result[8].31:=0;
   	End_If;
   	If UOWHF_Msg[10].[25] Then
   		UOWHF_Result[0]:=UOWHF_Result[0] + 1622696958+UOWHF_Add_c;
   		UOWHF_Add_c.0:=UOWHF_Result[0].31;
   		UOWHF_Result[0].31:=0;
   		UOWHF_Result[1]:=UOWHF_Result[1] + 592603911+UOWHF_Add_c;
   		UOWHF_Add_c.1:=UOWHF_Result[1].31;
   		UOWHF_Result[1].31:=0;
   		UOWHF_Result[2]:=UOWHF_Result[2] + 1448785737+UOWHF_Add_c;
   		UOWHF_Add_c.2:=UOWHF_Result[2].31;
   		UOWHF_Result[2].31:=0;
   		UOWHF_Result[3]:=UOWHF_Result[3] + 772462029+UOWHF_Add_c;
   		UOWHF_Add_c.3:=UOWHF_Result[3].31;
   		UOWHF_Result[3].31:=0;
   		UOWHF_Result[4]:=UOWHF_Result[4] + 265862720+UOWHF_Add_c;
   		UOWHF_Add_c.4:=UOWHF_Result[4].31;
   		UOWHF_Result[4].31:=0;
   		UOWHF_Result[5]:=UOWHF_Result[5] + 1600409915+UOWHF_Add_c;
   		UOWHF_Add_c.5:=UOWHF_Result[5].31;
   		UOWHF_Result[5].31:=0;
   		UOWHF_Result[6]:=UOWHF_Result[6] + 1971699096+UOWHF_Add_c;
   		UOWHF_Add_c.6:=UOWHF_Result[6].31;
   		UOWHF_Result[6].31:=0;
   		UOWHF_Result[7]:=UOWHF_Result[7] + 175967221+UOWHF_Add_c;
   		UOWHF_Add_c.7:=UOWHF_Result[7].31;
   		UOWHF_Result[7].31:=0;
   		UOWHF_Result[8]:=UOWHF_Result[8] + 2144844449+UOWHF_Add_c;
   		UOWHF_Add_c.8:=UOWHF_Result[8].31;
   		UOWHF_Result[8].31:=0;
   	End_If;
   	If UOWHF_Msg[10].[26] Then
   		UOWHF_Result[0]:=UOWHF_Result[0] + 1956517087+UOWHF_Add_c;
   		UOWHF_Add_c.0:=UOWHF_Result[0].31;
   		UOWHF_Result[0].31:=0;
   		UOWHF_Result[1]:=UOWHF_Result[1] + 662930096+UOWHF_Add_c;
   		UOWHF_Add_c.1:=UOWHF_Result[1].31;
   		UOWHF_Result[1].31:=0;
   		UOWHF_Result[2]:=UOWHF_Result[2] + 1272377109+UOWHF_Add_c;
   		UOWHF_Add_c.2:=UOWHF_Result[2].31;
   		UOWHF_Result[2].31:=0;
   		UOWHF_Result[3]:=UOWHF_Result[3] + 1761243004+UOWHF_Add_c;
   		UOWHF_Add_c.3:=UOWHF_Result[3].31;
   		UOWHF_Result[3].31:=0;
   		UOWHF_Result[4]:=UOWHF_Result[4] + 1810185770+UOWHF_Add_c;
   		UOWHF_Add_c.4:=UOWHF_Result[4].31;
   		UOWHF_Result[4].31:=0;
   		UOWHF_Result[5]:=UOWHF_Result[5] + 90808292+UOWHF_Add_c;
   		UOWHF_Add_c.5:=UOWHF_Result[5].31;
   		UOWHF_Result[5].31:=0;
   		UOWHF_Result[6]:=UOWHF_Result[6] + 282081916+UOWHF_Add_c;
   		UOWHF_Add_c.6:=UOWHF_Result[6].31;
   		UOWHF_Result[6].31:=0;
   		UOWHF_Result[7]:=UOWHF_Result[7] + 1588921715+UOWHF_Add_c;
   		UOWHF_Add_c.7:=UOWHF_Result[7].31;
   		UOWHF_Result[7].31:=0;
   		UOWHF_Result[8]:=UOWHF_Result[8] + 164466838+UOWHF_Add_c;
   		UOWHF_Add_c.8:=UOWHF_Result[8].31;
   		UOWHF_Result[8].31:=0;
   	End_If;
   	If UOWHF_Msg[10].[27] Then
   		UOWHF_Result[0]:=UOWHF_Result[0] + 447454653+UOWHF_Add_c;
   		UOWHF_Add_c.0:=UOWHF_Result[0].31;
   		UOWHF_Result[0].31:=0;
   		UOWHF_Result[1]:=UOWHF_Result[1] + 1088128821+UOWHF_Add_c;
   		UOWHF_Add_c.1:=UOWHF_Result[1].31;
   		UOWHF_Result[1].31:=0;
   		UOWHF_Result[2]:=UOWHF_Result[2] + 970436324+UOWHF_Add_c;
   		UOWHF_Add_c.2:=UOWHF_Result[2].31;
   		UOWHF_Result[2].31:=0;
   		UOWHF_Result[3]:=UOWHF_Result[3] + 486221453+UOWHF_Add_c;
   		UOWHF_Add_c.3:=UOWHF_Result[3].31;
   		UOWHF_Result[3].31:=0;
   		UOWHF_Result[4]:=UOWHF_Result[4] + 72190564+UOWHF_Add_c;
   		UOWHF_Add_c.4:=UOWHF_Result[4].31;
   		UOWHF_Result[4].31:=0;
   		UOWHF_Result[5]:=UOWHF_Result[5] + 1709022236+UOWHF_Add_c;
   		UOWHF_Add_c.5:=UOWHF_Result[5].31;
   		UOWHF_Result[5].31:=0;
   		UOWHF_Result[6]:=UOWHF_Result[6] + 575182992+UOWHF_Add_c;
   		UOWHF_Add_c.6:=UOWHF_Result[6].31;
   		UOWHF_Result[6].31:=0;
   		UOWHF_Result[7]:=UOWHF_Result[7] + 1495516910+UOWHF_Add_c;
   		UOWHF_Add_c.7:=UOWHF_Result[7].31;
   		UOWHF_Result[7].31:=0;
   		UOWHF_Result[8]:=UOWHF_Result[8] + 2069641147+UOWHF_Add_c;
   		UOWHF_Add_c.8:=UOWHF_Result[8].31;
   		UOWHF_Result[8].31:=0;
   	End_If;
   	If UOWHF_Msg[10].[28] Then
   		UOWHF_Result[0]:=UOWHF_Result[0] + 767079787+UOWHF_Add_c;
   		UOWHF_Add_c.0:=UOWHF_Result[0].31;
   		UOWHF_Result[0].31:=0;
   		UOWHF_Result[1]:=UOWHF_Result[1] + 544414095+UOWHF_Add_c;
   		UOWHF_Add_c.1:=UOWHF_Result[1].31;
   		UOWHF_Result[1].31:=0;
   		UOWHF_Result[2]:=UOWHF_Result[2] + 1962439250+UOWHF_Add_c;
   		UOWHF_Add_c.2:=UOWHF_Result[2].31;
   		UOWHF_Result[2].31:=0;
   		UOWHF_Result[3]:=UOWHF_Result[3] + 1977763716+UOWHF_Add_c;
   		UOWHF_Add_c.3:=UOWHF_Result[3].31;
   		UOWHF_Result[3].31:=0;
   		UOWHF_Result[4]:=UOWHF_Result[4] + 123363408+UOWHF_Add_c;
   		UOWHF_Add_c.4:=UOWHF_Result[4].31;
   		UOWHF_Result[4].31:=0;
   		UOWHF_Result[5]:=UOWHF_Result[5] + 288862386+UOWHF_Add_c;
   		UOWHF_Add_c.5:=UOWHF_Result[5].31;
   		UOWHF_Result[5].31:=0;
   		UOWHF_Result[6]:=UOWHF_Result[6] + 412670024+UOWHF_Add_c;
   		UOWHF_Add_c.6:=UOWHF_Result[6].31;
   		UOWHF_Result[6].31:=0;
   		UOWHF_Result[7]:=UOWHF_Result[7] + 641009862+UOWHF_Add_c;
   		UOWHF_Add_c.7:=UOWHF_Result[7].31;
   		UOWHF_Result[7].31:=0;
   		UOWHF_Result[8]:=UOWHF_Result[8] + 2110155119+UOWHF_Add_c;
   		UOWHF_Add_c.8:=UOWHF_Result[8].31;
   		UOWHF_Result[8].31:=0;
   	End_If;
   	If UOWHF_Msg[10].[29] Then
   		UOWHF_Result[0]:=UOWHF_Result[0] + 294706990+UOWHF_Add_c;
   		UOWHF_Add_c.0:=UOWHF_Result[0].31;
   		UOWHF_Result[0].31:=0;
   		UOWHF_Result[1]:=UOWHF_Result[1] + 2047620820+UOWHF_Add_c;
   		UOWHF_Add_c.1:=UOWHF_Result[1].31;
   		UOWHF_Result[1].31:=0;
   		UOWHF_Result[2]:=UOWHF_Result[2] + 1682273532+UOWHF_Add_c;
   		UOWHF_Add_c.2:=UOWHF_Result[2].31;
   		UOWHF_Result[2].31:=0;
   		UOWHF_Result[3]:=UOWHF_Result[3] + 450207604+UOWHF_Add_c;
   		UOWHF_Add_c.3:=UOWHF_Result[3].31;
   		UOWHF_Result[3].31:=0;
   		UOWHF_Result[4]:=UOWHF_Result[4] + 1417669551+UOWHF_Add_c;
   		UOWHF_Add_c.4:=UOWHF_Result[4].31;
   		UOWHF_Result[4].31:=0;
   		UOWHF_Result[5]:=UOWHF_Result[5] + 901079135+UOWHF_Add_c;
   		UOWHF_Add_c.5:=UOWHF_Result[5].31;
   		UOWHF_Result[5].31:=0;
   		UOWHF_Result[6]:=UOWHF_Result[6] + 1247347647+UOWHF_Add_c;
   		UOWHF_Add_c.6:=UOWHF_Result[6].31;
   		UOWHF_Result[6].31:=0;
   		UOWHF_Result[7]:=UOWHF_Result[7] + 472645253+UOWHF_Add_c;
   		UOWHF_Add_c.7:=UOWHF_Result[7].31;
   		UOWHF_Result[7].31:=0;
   		UOWHF_Result[8]:=UOWHF_Result[8] + 1986253441+UOWHF_Add_c;
   		UOWHF_Add_c.8:=UOWHF_Result[8].31;
   		UOWHF_Result[8].31:=0;
   	End_If;
   	If UOWHF_Msg[10].[30] Then
   		UOWHF_Result[0]:=UOWHF_Result[0] + 728151445+UOWHF_Add_c;